
   (* startup initialisation *)
   IF NOT #init OR #T = t#0s THEN
     #init := TRUE;
     #out := #K * #in;
   ELSE
     #out := #out + (#in * #K - #out) * DINT_TO_REAL(DWORD_TO_DINT(#tx) - DWORD_TO_DINT(#last)) / DINT_TO_REAL(T_CONV(#T)) * 1.0E-3;
     IF ABS(#out) < 1.0E-20 THEN #out := 0.0; END_IF;
   END_IF;
   #last := #tx;


   (*
   hm 1.1.2007 rev 1.1
     corrected error while startup value was not correct
     for very small time values real output would run out of range.

   hm 3.1.2007 rev 1.2
     corrected an error for falling edge failures.
     added output faktor K.

   hm 27. 2. 2007 rev 1.3
     output will be input during init for definitive startup condition.

   hm  15.9.2007 rev 1.4
     changed time() to T_PLC_US() for compatibilitxy resons
     increased internal accuracy to Microseconds instead of Milliseconds

   hm  23. oct 2007  rev 1.5
     added out := in to the init statements

   hm  30. nov 2007  rev 1.6
     changed out to be K * in during initialization

   hm  5. jan 2008 rev 1.7
     improved code for better performance

   hm  16. mar. 2008 rev 1.8
     added type conversion to avoid warning under codesys 3.0

   hm  14. jun. 2008 rev 1.9
     improved code

   hm  11. mar. 2009 rev 1.10
     real constants updated to new systax using dot

   hm  18. jan. 2011 rev 1.11
     avoid underrun of out
   *)
END_FUNCTION_BLOCK

FUNCTION_BLOCK "FT_PT2"   // FB163, SCL
TITLE = FT_PT2
{ S7_Optimized_Access := 'FALSE' }
AUTHOR : hugo
FAMILY : CTRL
NAME : PT2
VERSION : 1.5
// FT_PT2 is a 2nd grade filter with programmable times T, D and faktor K.
// 
// uses: INTEGRATE [FB237]
//       T_PLC_MS [FC64] 
//       STIME [FB64],IDB_STIME [DB64]
   VAR_INPUT
      in : Real;
      T : Time;
      D : Real;
      K : Real := 1.0e+0;
   END_VAR
   VAR_OUTPUT
      out : Real;
   END_VAR
   VAR
      init : Bool;
      int1 : "INTEGRATE";
      int2 : "INTEGRATE";
      tn : Real;
      I1 : Real;
      I2 : Real;
      tn2 : Real;
   END_VAR
BEGIN


   (* startup initialisation *)
   IF NOT #init OR #T = T#0s THEN
       #init := TRUE;
       #out := #K * #in;
       #I2 := #out;
   ELSE
       #tn := DINT_TO_REAL(T_CONV(#T)) * 1.0E-3;
       #tn2 := #tn * #tn;
       #int1(X := #in * #K / #tn2 - #I1 * 0.5 * #D / #tn - #I2 / #tn2, Y := #I1);
       #int2(X := #I1,Y := #I2);
       #out := #I2;
   END_IF;


   (* revision history

   15.1.2007 hm        rev 1.1
       changed formula to new more acurate formula

   hm 15.9.2007        rev 1.2
       deleted unused code for init system time reading tx 

   hm  30.11.2007  rev 1.3
       changed out to be K * in during initialization
       avoind divide by 0 if tn = 0

   hm  3. nov. 2008    rev 1.4
       optimized code and fixed a problem with init

   hm  11. mar. 2009   rev 1.5
       real constants updated to new systax using dot

   *)
END_FUNCTION_BLOCK

FUNCTION_BLOCK "FT_TN16"   // FB164, SCL
TITLE = FT_TN16
{ S7_Optimized_Access := 'FALSE' }
AUTHOR : hugo
FAMILY : CTRL
NAME : TN16
VERSION : 1.1
// FT_TN16 is delay function, it will delay a signal by a specified time : T and will store 16 values of in before they are put thru to out.
// for higher OR lower resolution please use FT_TN8 OR FT_TN64 instead.
// 
// uses: T_PLC_MS [FC64]
//       STIME [FB64],IDB_STIME [DB64]
   VAR_INPUT
      in : Real;
      T : Time;
   END_VAR
   VAR_OUTPUT
      out : Real;
      trig : Bool;
   END_VAR
   VAR
      length : Int := 16;
      X : Array[0..15] of Real;
      cnt : Int;
      last : Time;
      tx : Time;
      init : Bool;
   END_VAR
BEGIN


     (* read system time *)
     #tx := T_CONV(DWORD_TO_DINT("T_PLC_MS"()));

     #trig := FALSE;
     IF NOT #init THEN
       #X[#cnt] := #in;
       #init := TRUE;
       #last := #tx;
     ELSIF #tx - #last >= #T / #length THEN
       IF #cnt = #length - 1 THEN #cnt := 0; ELSE #cnt := #cnt + 1; END_IF;
       #out := #X[#cnt];
       #X[#cnt] := #in;
       #last := #tx;
       #trig := TRUE;
     END_IF;

   (* revision history
   hm    1. jan 2007    rev 1.0
     original version

   hm    16. sep 2007  rev 1.1
     changes time() to T_plc_ms() for compatibility reasons

   *)
END_FUNCTION_BLOCK

FUNCTION_BLOCK "FT_TN64"   // FB165, SCL
TITLE = FT_TN64
{ S7_Optimized_Access := 'FALSE' }
AUTHOR : hugo
FAMILY : CTRL
NAME : TN64
VERSION : 1.1
// FT_TN64 is delay function, it will delay a signal by a specified time : T and will store 64 values of in before they are put thru to out.
// if lower resolution is needed, pls use FT_TN8 or FT_TN16 instead.
// 
// uses: T_PLC_MS [FC64]
//       STIME [FB64],IDB_STIME [DB64]
   VAR_INPUT
      in : Real;
      T : Time;
   END_VAR
   VAR_OUTPUT
      out : Real;
      trig : Bool;
   END_VAR
   VAR
      length : Int := 64;
      X : Array[0..63] of Real;
      cnt : Int;
      last : Time;
      tx : Time;
      init : Bool;
   END_VAR
BEGIN


     (* read system time *)
     #tx := T_CONV(DWORD_TO_DINT("T_PLC_MS"()));

     #trig := FALSE;
     IF NOT #init THEN
       #X[#cnt] := #in;
       #init := TRUE;
       #last := #tx;
     ELSIF #tx - #last >= #T / #length THEN
       IF #cnt = #length - 1 THEN #cnt := 0; ELSE #cnt := #cnt + 1; END_IF;
       #out := #X[#cnt];
       #X[#cnt] := #in;
       #last := #tx;
       #trig := TRUE;
     END_IF;

   (* revision history
   hm    1. jan 2007    rev 1.0
     original version

   hm    16. sep 2007  rev 1.1
     changes time() to T_plc_ms() for compatibility reasons

   *)
END_FUNCTION_BLOCK

FUNCTION_BLOCK "FT_TN8"   // FB166, SCL
TITLE = FT_TN8
{ S7_Optimized_Access := 'FALSE' }
AUTHOR : hugo
FAMILY : CTRL
NAME : TN8
VERSION : 1.1
// FT_TN8 is delay function, it will delay a signal by a specified time : T and will store 8 values of in before they are put thru to out.
// if higher resolution is needed, pls use FT_TN16 or FT_TN64 instead.
// 
// uses: T_PLC_MS [FC64]
//       STIME [FB64],IDB_STIME [DB64]
   VAR_INPUT
      in : Real;
      T : Time;
   END_VAR
   VAR_OUTPUT
      out : Real;
      trig : Bool;
   END_VAR
   VAR
      length : Int := 8;
      X : Array[0..7] of Real;
      cnt : Int;
      last : Time;
      tx : Time;
      init : Bool;
   END_VAR
BEGIN


     #tx := T_CONV(DWORD_TO_DINT("T_PLC_MS"()));
     #trig := FALSE;
     IF NOT #init THEN
       #X[#cnt] := #in;
       #init := TRUE;
       #last := #tx;
     ELSIF #tx - #last >= #T / #length THEN
       IF #cnt = #length - 1 THEN #cnt := 0; ELSE #cnt := #cnt + 1; END_IF;
       #out := #X[#cnt];
       #X[#cnt] := #in;
       #last := #tx;
       #trig := TRUE;
     END_IF;

   (* revision history
   hm    1. jan 2007    rev 1.0
     original version

   hm    16. sep 2007  rev 1.1
     changes time() to T_plc_ms() for compatibility reasons

   *)
END_FUNCTION_BLOCK

FUNCTION_BLOCK "HYST"   // FB167, SCL
TITLE = HYST
{ S7_Optimized_Access := 'FALSE' }
AUTHOR : hugo
FAMILY : CTRL
NAME : HYST
VERSION : 1.0
// This Hystereses function has two modes:
// 1. if on > off then Q will be switched high when in > on and switched low when in < off.
// 2. if on < off then Q will be switched high when in < on and switched low when in > off.
// the output win will be high when in is between low and high.
   VAR_INPUT
      In : Real;
      ON : Real;
      OFF : Real;
   END_VAR
   VAR_OUTPUT
      Q : Bool;
      win : Bool;
   END_VAR
BEGIN


   IF #ON >= #OFF THEN
       IF #In < #OFF THEN
           #Q := FALSE;
           #win := FALSE;
       ELSIF  #In > #ON THEN
           #Q := TRUE;
           #win := FALSE;
       ELSE
           #win := TRUE;
       END_IF;
   ELSE
       IF #In > #OFF THEN
           #Q := FALSE;
           #win := FALSE;
       ELSIF  #In < #ON THEN
           #Q := TRUE;
           #win := FALSE;
       ELSE
           #win := TRUE;
       END_IF;
   END_IF;


   (* revision history
   hm      2.  jun 2008    rev 1.0
       original version

   *)
END_FUNCTION_BLOCK

FUNCTION_BLOCK "HYST_1"   // FB168, SCL
TITLE = HYST_1
{ S7_Optimized_Access := 'FALSE' }
AUTHOR : hugo
FAMILY : CTRL
NAME : HYST_1
VERSION : 1.1
// this hysteresis function switches the output high if the input signal reaches obove high and will switch to low when the input falls back below low value.
// a separate output mid is set if the input stays between low and high value.
   VAR_INPUT
      In : Real;
      high : Real;
      low : Real;
   END_VAR
   VAR_OUTPUT
      Q : Bool;
      win : Bool;
   END_VAR
BEGIN


   IF #In < #low THEN
       #Q := FALSE;
       #win := FALSE;
   ELSIF #In > #high THEN
       #Q := TRUE;
       #win := FALSE;
   ELSE
       #win := TRUE;
   END_IF;

   (* code used for rev 1.0
   IF Q THEN
       IF in < low THEN q := FALSE; END_IF;
   ELSE
       IF in > high THEN q := TRUE; END_IF;
   END_IF;
   win := in > low AND in < high;
   *)


   (* revision history
   hm      4.  aug. 2006   rev 1.0
       original version

   hm      2. jun. 2008    rev 1.1
       improved performance
   *)
END_FUNCTION_BLOCK

FUNCTION_BLOCK "HYST_2"   // FB169, SCL
TITLE = HYST_2
{ S7_Optimized_Access := 'FALSE' }
AUTHOR : oscat
FAMILY : CTRL
NAME : HYST_2
VERSION : 1.2
// this hysteresis function switches the output high if the input signal reaches obove val + hys/2 and will switch to low when the input falls back below val - hys/2 value.
// a separate output mid is set if the input stays between low and high value.
   VAR_INPUT
      IN : Real;
      VAL : Real;
      HYS : Real;
   END_VAR
   VAR_OUTPUT
      Q : Bool;
      WIN : Bool;
   END_VAR
   VAR
      tmp : Real;
   END_VAR
BEGIN


   #tmp := #VAL - #HYS * 0.5;
   IF #IN < #tmp THEN
       #Q := FALSE;
       #WIN := FALSE;
   ELSIF #IN > #tmp + #HYS THEN
       #Q := TRUE;
       #WIN := FALSE;
   ELSE
       #WIN := TRUE;
   END_IF;

   (* code used for 1.2 and before
   X := hys * 0.5;
   IF Q THEN
       IF in < val - x THEN q := FALSE; END_IF;
   ELSE
       IF in > val + x THEN q := TRUE; END_IF;
   END_IF;
   win := in > val - x AND in < val + x;
   *)

   (* revision history
   hm      4. aug 2006 rev 1.0
       original version

   hm      5. jan 2008 rev 1.1
       improved code for better performance

   hm      2. jun. 2008    rev 1.2
       improved performance
   *)
END_FUNCTION_BLOCK

FUNCTION_BLOCK "HYST_3"   // FB170, SCL
TITLE = HYST_3
{ S7_Optimized_Access := 'FALSE' }
AUTHOR : oscat
FAMILY : CTRL
NAME : HYST_3
VERSION : 1.2
// this is a double hysteresis function. Out1 follows a hysteresis function defined by val1and hyst, while out 2 follows val2 and hyst.
// if the input signal is between the two hysteresis switches (val1 and val2) then non of the outputs is active.
   VAR_INPUT
      in : Real;
      hyst : Real;
      val1 : Real;
      val2 : Real;
   END_VAR
   VAR_OUTPUT
      Q1 : Bool;
      Q2 : Bool;
   END_VAR
   VAR
      X : Real;
   END_VAR
BEGIN


     #X := #hyst * 0.5;

     IF #in < #val1 - #X THEN
         #Q1 := TRUE;
     ELSIF #in > #val1 + #X THEN
         #Q1 := FALSE;
     END_IF;
     IF #in < #val2 - #X THEN
         #Q2 := FALSE;
     ELSIF #in > #val2 + #X THEN
         #Q2 := TRUE;
     END_IF;

   (* revision history
   hm  22. jan 2007  rev 1.0
     original version

   hm  27. dec 2007  rev 1.1
     changed code for better performance

   hm  5. jan 2008   rev 1.2
     further performance iprovements

   *)
END_FUNCTION_BLOCK

FUNCTION_BLOCK "INTEGRATE"   // FB237, SCL
TITLE = INTEGRATE
{ S7_Optimized_Access := 'FALSE' }
AUTHOR : hugo
FAMILY : CTRL
NAME : INTEGR
VERSION : 1.0
// integrate is a plain integrator with I/O for out.
// 
// uses: T_PLC_MS [FC64]
//       STIME [FB64],IDB_STIME [DB64]
   VAR_INPUT
      "E" : Bool := TRUE;
      X : Real;
      K : Real := 1.0e+0;
   END_VAR
   VAR_IN_OUT
      Y : Real;
   END_VAR
   VAR
      X_last : Real;
      init : Bool;
      last : DWord;
      tx : DWord;
   END_VAR
   VAR_TEMP
      TOP_SI : Struct
         EV_CLASS : Byte;
         EV_NUM : Byte;
         PRIORITY : Byte;
         NUM : Byte;
         TYP2_3 : Byte;
         TYP1 : Byte;
         ZI1 : Word;
         ZI2_3 : DWord;
      END_STRUCT;
      START_UP_SI : Struct
         EV_CLASS : Byte;
         EV_NUM : Byte;
         PRIORITY : Byte;
         NUM : Byte;
         TYP2_3 : Byte;
         TYP1 : Byte;
         ZI1 : Word;
         ZI2_3 : DWord;
      END_STRUCT;
      ERR : Int;
   END_VAR
BEGIN


   (* read actual startup info *)
   (* OB1_SCAN_1  BYTE  -  B#16#01: Abschluss des Neustarts (Warmstarts)
                        -  B#16#02: Abschluss des Wiederanlaufs
                        -  B#16#03: Abschluss des freien Zyklus
                        -  B#16#04: Abschluss des Kaltstarts
                        -  B#16#05: Erster OB 1-Zyklus der neuen Master-CPU nach 
                                    Master-Reserve-Umschaltung und STOP des 
                                    bisherigen Masters *)

   #ERR := RD_SINFO (TOP_SI => #TOP_SI, START_UP_SI => #START_UP_SI);

   (* reset last_time on system startup *)
   IF #TOP_SI.EV_NUM = 1 OR #TOP_SI.EV_NUM = 2 OR #TOP_SI.EV_NUM = 4 THEN 
       #init := FALSE;
   END_IF;

   (*read system time *)
   #tx := "T_PLC_MS"();

   IF NOT #init THEN
       #init := TRUE;
       #X_last := #X;
   ELSIF #"E" THEN
       #Y := (#X + #X_last) * 0.5E-3 * DINT_TO_REAL(DWORD_TO_DINT(#tx)-DWORD_TO_DINT(#last)) * #K + #Y;
       #X_last := #X;
   END_IF;
   #last := #tx;


   (*
   hm  3. nov. 2008    rev 1.0
   original version

   *)
END_FUNCTION_BLOCK

FUNCTION "T_PLC_MS" : DWord   // FC64, SCL
TITLE = T_PLC_MS
{ S7_Optimized_Access := 'FALSE' }
AUTHOR : hugo
FAMILY : MEASURE
NAME : T_PLC_MS
VERSION : 1.2
// T_PLC_MS reads the internal PLC timer and return the time, it has the advantage to be able to set a debug mode 
// and speed up the counter to test the plc timer overrun which occurs every 50 days respectively 25 days at siemens S7
// this routine also allows to correct the behavior of s7 where the internal plc counter will not count all 32 bits.
// 
// uses: STIME [FB64],IDB_STIME [DB64]
BEGIN


   "IDB_STIME"(); 
   #T_PLC_MS := "IDB_STIME".tx; 
   (* hier muss die korrektur für step7 stattfinden
   plctime muss den vollen wertebereich von time ausnutzen:
   wenn bei step7 time -24tage bis plus 24 tage ist dann muss der timer auch beim überlauf auf -24tage springen 
   und auf keinen fall auf 0 !!!!
   für siemens muss ein weiterer fb im main eingebunden werden der sicherstellt das alle 32 bits durchgezählt werden.
   es kann nur ein fb sein den er muss sich das oberste (32te) bit merken.
   oder etwa spring s7 bei überlauf auf -24 tage????? dann wäre keine korrektur nötig.
   *)
   IF "debug" THEN
       #T_PLC_MS := DINT_TO_DWORD((DWORD_TO_DINT(SHL(IN:=#T_PLC_MS,N:="N") OR SHL(IN:=DWORD#1,N:="N"))-1) + DWORD_TO_DINT("offset_1"));
   END_IF;


   (* revision history
   hm  14.9.2007   rev 1.0
       original version

   hm  12. nov 2007    rev 1.1
       added temporaray variable tx because some compilers could not handle time() as an argument

   hm  16. nov. 2008   rev 1.2
       initialized constants with 0 for compatibility reasons
   *)
END_FUNCTION

FUNCTION "T_PLC_US" : DWord   // FC65, SCL
TITLE = T_PLC_US
{ S7_Optimized_Access := 'FALSE' }
AUTHOR : hugo
FAMILY : MEASURE
NAME : T_PLC_US
VERSION : 1.2
// T_PLC_US reads the internal PLC timer and return the time, it has the advantage to be able to set a debug mode 
// and speed up the counter to test the plc timer overrun which occurs every 50 days respectively 25 days at siemens S7
// this routine also allows to correct the behavior of s7 where the internal plc counter will not count all 32 bits.
// 
// uses: STIME [FB64],IDB_STIME [DB64]
BEGIN


   "IDB_STIME"(); 
   #T_PLC_US := DINT_TO_DWORD(DWORD_TO_DINT("IDB_STIME".tx) * 1000); 
   (* hier muss die korrektur für step7 stattfinden
   plctime muss den vollen wertebereich von time ausnutzen:
   wenn bei step7 time -24tage bis plus 24 tage ist dann muss der timer auch beim überlauf auf -24tage springen 
   und auf keinen fall auf 0 !!!!
   für siemens muss ein weiterer fb im main eingebunden werden der sicherstellt das alle 32 bits durchgezählt werden.
   es kann nur ein fb sein den er muss sich das oberste (32te) bit merken.
   oder etwa spring s7 bei überlauf auf -24 tage????? dann wäre keine korrektur nötig.
   *)
   IF "debug" THEN
       #T_PLC_US := DINT_TO_DWORD((DWORD_TO_DINT(SHL(IN:=#T_PLC_US,N:="N") OR SHL(IN:=DWORD#1,N:="N"))-1) + DWORD_TO_DINT("offset_1"));
   END_IF;


   (* revision history
   hm  14.9.2007   rev 1.0
       original version

   hm  12. nov 2007    rev 1.1
       added temporaray variable tx because some compilers could not handle time() as an argument

   hm  16. nov. 2008   rev 1.2
       initialized constants with 0 for compatibility reasons

   *)
END_FUNCTION

FUNCTION "R2_ADD" : "REAL2"   // FC144, SCL
TITLE = R2_ADD
{ S7_Optimized_Access := 'FALSE' }
AUTHOR : hugo
FAMILY : R2
NAME : ADD
VERSION : 1.0
// R2_add adds a real to a double real which extends the accuracy of a real to twice as many digits
//  
// uses: REAL2 [UDT11]
   VAR_INPUT
      X : "REAL2";
      Y : Real;
   END_VAR
   VAR_TEMP
      temp : Real;
      tR2_ADD : "REAL2";
   END_VAR
BEGIN


   #temp := #X.RX;
   #tR2_ADD.RX := #Y + #X.R1 + #X.RX;
   #tR2_ADD.R1 := #temp - #tR2_ADD.RX + #Y + #X.R1;

   #R2_ADD := #tR2_ADD;

   (* revision history
   hm      20.3.2008   rev 1.0
       original version

   *)
END_FUNCTION

FUNCTION "R2_SET" : "REAL2"   // FC147, SCL
TITLE = R2_SET
{ S7_Optimized_Access := 'FALSE' }
AUTHOR : hugo
FAMILY : R2
NAME : SET
VERSION : 1.1
// R2_set sets a double precision real to a single real value.
// 
// uses: REAL2 [UDT11]
   VAR_INPUT
      X : Real;
   END_VAR
   VAR_TEMP
      tR2_SET : "REAL2";
   END_VAR
BEGIN


   #tR2_SET.RX := #X;
   #tR2_SET.R1 := 0.0;

   #R2_SET := #tR2_SET;


   (* revision history
   hm  2. jun. 2008    rev 1.0
       original version

   hm  10. mar. 2009   rev 1.1
       real constants updated to new systax using dot

   *)
END_FUNCTION

FUNCTION "MULTIME" : Time   // FC203, SCL
TITLE = MULTIME
{ S7_Optimized_Access := 'FALSE' }
AUTHOR : hugo
FAMILY : TIDT
NAME : MULTIME
VERSION : 1.1
// multiplies a time by a real number and returns a time
   VAR_INPUT
      t : Time;
      "M" : Real;
   END_VAR
BEGIN


     #MULTIME := T_CONV(REAL_TO_DINT(DINT_TO_REAL(T_CONV(#t))*#"M"));

   (* revision history
   hm      2. oct 2006 rev 1.0
       original version

   hm      14. mar 2008    rev 1.1
       rounded the result after the last digit

   *)
END_FUNCTION

FUNCTION "CTRL_IN" : Real   // FC363, SCL
TITLE = CTRL_IN
{ S7_Optimized_Access := 'FALSE' }
AUTHOR : hugo
FAMILY : CTRL
NAME : CTRL_IN
VERSION : 1.0
// uses: DEAD_ZONE [FC365]
   VAR_INPUT
      SET_POINT : Real;
      ACTUAL : Real;
      NOISE : Real;
   END_VAR
BEGIN


   (* calculate the process error DIFF *)
   #CTRL_IN := "DEAD_ZONE"(X:=#SET_POINT - #ACTUAL,L:=#NOISE);


   (* revision history
   hm  2. jun. 2008    rev 1.0
       original version

   *)
END_FUNCTION

FUNCTION "DEAD_BAND" : Real   // FC364, SCL
TITLE = DEAD_BAND
{ S7_Optimized_Access := 'FALSE' }
AUTHOR : hugo
FAMILY : CTRL
NAME : DEADBAND
VERSION : 1.2
// DEAD_BAND ist eine lineare Übertragungsfunktion mit Totzone. Die Funktion verschiebt den positiven Teil der Kurve um +L und den negativen Teil der Kurve um -L.
// DEAD_BAND = X - L wenn X > L)
// DEAD_BAND = X + L wenn X < -L
// DEAD_BAND = 0 wenn Abs(X) <= L
   VAR_INPUT
      X : Real;
      L : Real;
   END_VAR
BEGIN


     IF #X > #L THEN
       #DEAD_BAND := #X - #L;
     ELSIF #X < -#L THEN
       #DEAD_BAND := #X + #L;
     ELSE
       #DEAD_BAND := 0.0;
     END_IF;


   (* revision history
   hm  2. nov. 2007  rev 1.0
     original version

   hm  14. jun. 2008 rev 1.1
     improved performance

   hm  18. jan. 2011 rev 1.2
     assign 0 before return
   *)
END_FUNCTION

FUNCTION "DEAD_ZONE" : Real   // FC365, SCL
TITLE = DEAD_ZONE
{ S7_Optimized_Access := 'FALSE' }
AUTHOR : hugo
FAMILY : CTRL
NAME : DEADZONE
VERSION : 1.2
// dead_zone2 is a linear transfer function which follows a linear function except for x is close to 0.
// Y = X if abs(x) > L otherwise its 0.
   VAR_INPUT
      X : Real;
      L : Real;
   END_VAR
BEGIN


   IF ABS(#X) > #L THEN
       #DEAD_ZONE := #X;
   ELSE
       #DEAD_ZONE := 0.0;
   END_IF;


   (* revision history
   hm  12. feb. 2007   rev 1.0
       original version

   hm  14. jun. 2008   rev 1.1
       improved performance

   hm  11. mar. 2009   rev 1.2
       real constants updated to new systax using dot

   *)
END_FUNCTION

FUNCTION "BAND_B" : Byte   // FC410, SCL
TITLE = BAND_B
{ S7_Optimized_Access := 'FALSE' }
AUTHOR : hugo
FAMILY : CTRL
NAME : BAND_B
VERSION : 1.0
// BAND_B will limit X to B <= X <= 255-B. while X < B the resulkt will be 0 and while X > 255-B the output will be 255
// otherwise the result = X.
   VAR_INPUT
      X : Byte;
      "B" : Byte;
   END_VAR
BEGIN


   IF BYTE_TO_INT(#X) < BYTE_TO_INT(#"B") THEN
       #BAND_B := 0;
   ELSIF BYTE_TO_INT(#X) > BYTE_TO_INT(BYTE#255) - BYTE_TO_INT(#"B") THEN
       #BAND_B := 255;
   ELSE
       #BAND_B := #X;
   END_IF;



   (* revision history
   hm  21. nov. 2008   rev 1.0
       original version

   *)
END_FUNCTION

// ===== PLC "Engineering conversion"  Unspecific CPU S7 300 =====

VAR_GLOBAL CONSTANT   // PLC tag table "STEP7 classic symbols"
   "#T0" : Real := -2.731500E+002;   // MigChange: -273.15 OriginalComment: absoluter Nullpunkt in °C
   "PI2" : Real := 6.28318530717958647692528676655900576;   // PI * 2
END_VAR

DATA_BLOCK "LANGUAGE"   // DB4
TITLE = LANGUAGE
{ S7_Optimized_Access := 'FALSE' }
AUTHOR : oscat
FAMILY : CONSTANT
NAME : DBLANG
VERSION : 1.2
   VAR
      DEFAULT : Int := 1;   // 1=english, 2=german, 3=french
      LMAX : Int := 3;
      WEEKDAYS : Array[1..3, 1..7] of String[10];
      WEEKDAYS2 : Array[1..3, 1..7] of String[2];
      MONTHS : Array[1..3, 1..12] of String[10];
      MONTHS3 : Array[1..3, 1..12] of String[3];
      DIRS : Array[1..3, 0..15] of String[3];
   END_VAR
BEGIN
   WEEKDAYS[1,1] := 'Monday';
   WEEKDAYS[1,2] := 'Tuesday';
   WEEKDAYS[1,3] := 'Wednesday';
   WEEKDAYS[1,4] := 'Thursday';
   WEEKDAYS[1,5] := 'Friday';
   WEEKDAYS[1,6] := 'Saturday';
   WEEKDAYS[1,7] := 'Sunday';
   WEEKDAYS[2,1] := 'Montag';
   WEEKDAYS[2,2] := 'Dienstag';
   WEEKDAYS[2,3] := 'Mittwoch';
   WEEKDAYS[2,4] := 'Donnerstag';
   WEEKDAYS[2,5] := 'Freitag';
   WEEKDAYS[2,6] := 'Samstag';
   WEEKDAYS[2,7] := 'Sonntag';
   WEEKDAYS[3,1] := 'Lundi';
   WEEKDAYS[3,2] := 'Mardi';
   WEEKDAYS[3,3] := 'Mercredi';
   WEEKDAYS[3,4] := 'Jeudi';
   WEEKDAYS[3,5] := 'Vendredi';
   WEEKDAYS[3,6] := 'Samedi';
   WEEKDAYS[3,7] := 'Dimanche';
   WEEKDAYS2[1,1] := 'Mo';
   WEEKDAYS2[1,2] := 'Tu';
   WEEKDAYS2[1,3] := 'We';
   WEEKDAYS2[1,4] := 'Th';
   WEEKDAYS2[1,5] := 'Fr';
   WEEKDAYS2[1,6] := 'Sa';
   WEEKDAYS2[1,7] := 'Su';
   WEEKDAYS2[2,1] := 'Mo';
   WEEKDAYS2[2,2] := 'Di';
   WEEKDAYS2[2,3] := 'Mi';
   WEEKDAYS2[2,4] := 'Do';
   WEEKDAYS2[2,5] := 'Fr';
   WEEKDAYS2[2,6] := 'Sa';
   WEEKDAYS2[2,7] := 'So';
   WEEKDAYS2[3,1] := 'Lu';
   WEEKDAYS2[3,2] := 'Ma';
   WEEKDAYS2[3,3] := 'Me';
   WEEKDAYS2[3,4] := 'Je';
   WEEKDAYS2[3,5] := 'Ve';
   WEEKDAYS2[3,6] := 'Sa';
   WEEKDAYS2[3,7] := 'Di';
   MONTHS[1,1] := 'January';
   MONTHS[1,2] := 'February';
   MONTHS[1,3] := 'March';
   MONTHS[1,4] := 'April';
   MONTHS[1,5] := 'May';
   MONTHS[1,6] := 'June';
   MONTHS[1,7] := 'July';
   MONTHS[1,8] := 'August';
   MONTHS[1,9] := 'September';
   MONTHS[1,10] := 'October';
   MONTHS[1,11] := 'November';
   MONTHS[1,12] := 'December';
   MONTHS[2,1] := 'Januar';
   MONTHS[2,2] := 'Februar';
   MONTHS[2,3] := 'März';
   MONTHS[2,4] := 'April';
   MONTHS[2,5] := 'Mai';
   MONTHS[2,6] := 'Juni';
   MONTHS[2,7] := 'Juli';
   MONTHS[2,8] := 'August';
   MONTHS[2,9] := 'September';
   MONTHS[2,10] := 'Oktober';
   MONTHS[2,11] := 'November';
   MONTHS[2,12] := 'Dezember';
   MONTHS[3,1] := 'Janvier';
   MONTHS[3,2] := 'Février';
   MONTHS[3,3] := 'mars';
   MONTHS[3,4] := 'Avril';
   MONTHS[3,5] := 'Mai';
   MONTHS[3,6] := 'Juin';
   MONTHS[3,7] := 'Juillet';
   MONTHS[3,8] := 'Août';
   MONTHS[3,9] := 'Septembre';
   MONTHS[3,10] := 'Octobre';
   MONTHS[3,11] := 'Novembre';
   MONTHS[3,12] := 'Decembre';
   MONTHS3[1,1] := 'Jan';
   MONTHS3[1,2] := 'Feb';
   MONTHS3[1,3] := 'Mar';
   MONTHS3[1,4] := 'Apr';
   MONTHS3[1,5] := 'May';
   MONTHS3[1,6] := 'Jun';
   MONTHS3[1,7] := 'Jul';
   MONTHS3[1,8] := 'Aug';
   MONTHS3[1,9] := 'Sep';
   MONTHS3[1,10] := 'Oct';
   MONTHS3[1,11] := 'Nov';
   MONTHS3[1,12] := 'Dec';
   MONTHS3[2,1] := 'Jan';
   MONTHS3[2,2] := 'Feb';
   MONTHS3[2,3] := 'Mrz';
   MONTHS3[2,4] := 'Apr';
   MONTHS3[2,5] := 'Mai';
   MONTHS3[2,6] := 'Jun';
   MONTHS3[2,7] := 'Jul';
   MONTHS3[2,8] := 'Aug';
   MONTHS3[2,9] := 'Sep';
   MONTHS3[2,10] := 'Okt';
   MONTHS3[2,11] := 'Nov';
   MONTHS3[2,12] := 'Dez';
   MONTHS3[3,1] := 'Jan';
   MONTHS3[3,2] := 'Fev';
   MONTHS3[3,3] := 'Mar';
   MONTHS3[3,4] := 'Avr';
   MONTHS3[3,5] := 'Mai';
   MONTHS3[3,6] := 'Jun';
   MONTHS3[3,7] := 'Jul';
   MONTHS3[3,8] := 'Aou';
   MONTHS3[3,9] := 'Sep';
   MONTHS3[3,10] := 'Oct';
   MONTHS3[3,11] := 'Nov';
   MONTHS3[3,12] := 'Dec';
   DIRS[1,0] := 'N';
   DIRS[1,1] := 'NNE';
   DIRS[1,2] := 'NE';
   DIRS[1,3] := 'ENE';
   DIRS[1,4] := 'E';
   DIRS[1,5] := 'ESE';
   DIRS[1,6] := 'SE';
   DIRS[1,7] := 'SSE';
   DIRS[1,8] := 'S';
   DIRS[1,9] := 'SSW';
   DIRS[1,10] := 'SW';
   DIRS[1,11] := 'WSW';
   DIRS[1,12] := 'W';
   DIRS[1,13] := 'WNW';
   DIRS[1,14] := 'NW';
   DIRS[1,15] := 'NNW';
   DIRS[2,0] := 'N';
   DIRS[2,1] := 'NNO';
   DIRS[2,2] := 'NO';
   DIRS[2,3] := 'ONO';
   DIRS[2,4] := 'O';
   DIRS[2,5] := 'OSO';
   DIRS[2,6] := 'SO';
   DIRS[2,7] := 'SSO';
   DIRS[2,8] := 'S';
   DIRS[2,9] := 'SSW';
   DIRS[2,10] := 'SW';
   DIRS[2,11] := 'WSW';
   DIRS[2,12] := 'W';
   DIRS[2,13] := 'WNW';
   DIRS[2,14] := 'NW';
   DIRS[2,15] := 'NNW';
   DIRS[3,0] := 'N';
   DIRS[3,1] := 'NNO';
   DIRS[3,2] := 'NO';
   DIRS[3,3] := 'ONO';
   DIRS[3,4] := 'O';
   DIRS[3,5] := 'OSO';
   DIRS[3,6] := 'SO';
   DIRS[3,7] := 'SSO';
   DIRS[3,8] := 'S';
   DIRS[3,9] := 'SSW';
   DIRS[3,10] := 'SW';
   DIRS[3,11] := 'WSW';
   DIRS[3,12] := 'W';
   DIRS[3,13] := 'WNW';
   DIRS[3,14] := 'NW';
   DIRS[3,15] := 'NNW';
END_DATA_BLOCK

FUNCTION_BLOCK "ASTRO"   // FB136, SCL
TITLE = ASTRO
{ S7_Optimized_Access := 'FALSE' }
AUTHOR : oscat
FAMILY : CONVERT
NAME : ASTRO
VERSION : 1.1
// this function converts different length units
// any unused input can simply be left open.
// different inputs connected at the same time will be added up.
   VAR_INPUT
      "m" : Real;
      AE : Real;
      PC : Real;
      LJ : Real;
   END_VAR
   VAR_OUTPUT
      Ym : Real;
      YAE : Real;
      YPC : Real;
      YLJ : Real;
   END_VAR
BEGIN


   #YAE :=  #AE
           + #"m" * 6.6845871535E-012
           + #PC * 206265.0
           + #LJ * 63240.0;
   #Ym := #YAE * 149.597870E9;
   #YPC := #YAE * 4.8481322570E-006;
   #YLJ := #YAE * 1.5812776724E-005;


   (*
   Länge Meter m SI-Basiseinheit
   Astronomische Einheit* AE 1 AE = 149,597 870 · E9 m
   Parsec pc 1 pc = 206265 AE = 30,857 · E15 m
   Lichtjahr Lj 1 Lj = 9,460 530 · E15 m = 63240 AE = 0,306 59 pc
   Ångström Å 1 Å = E–l0 m
   typograph. Punkt p 1 p = 0,376 065 mm • im Druckereigewerbe
   inch** in 1 in = 2,54 · E–2 m = 25,4 mm***
   foot ft 1 ft = 0,3048 m = 30,48 cm
   yard yd 1 yd = 0,9144 m
   mile mile 1 mile = 1609,344 m
   Internat. Seemeile sm 1 sm = 1852 m
   Fathom fm 1 fm = 1,829 m • in der Seeschifffahrt
   *)

   (* revision history

   hm  27. mar. 2007   rev 1.0
       original version

   hm  11. mar. 2009   rev 1.1
       improved code

   *)
END_FUNCTION_BLOCK

FUNCTION_BLOCK "ENERGY"   // FB137, SCL
TITLE = ENERGY
{ S7_Optimized_Access := 'FALSE' }
AUTHOR : hugo
FAMILY : CONVERT
NAME : ENERGY
VERSION : 1.2
// this function converts different energy units
// any unused input can simply be left open.
// different inputs connected at the same time will be added up.
   VAR_INPUT
      J : Real;
      C : Real;
      Wh : Real;
   END_VAR
   VAR_OUTPUT
      YJ : Real;
      YC : Real;
      YWh : Real;
   END_VAR
BEGIN


   #YJ := #J + #Wh * 3600.0 + #C * 4.1868;
   #YC := #YJ * 0.238845896627496;
   #YWh := #YJ * 2.7777777778E-004;


   (*
   Arbeit, Energie, Joule* J 1 J = 1 N · m = 1 W · s = (1/3,6) E–6 kW · h = 1 kg · m2/s2
   Wärmemenge Kilowattstunde kW · h 1 kW · h = 3,6 MJ = 860 kcal
   Elektronvolt eV 1 eV = 160,218 92 E–21 J
   Erg erg 1 erg = 1E–7 J
   Kalorie cal 1 cal = 4,1868 J = 1,163 E–3 W · h
   Therm therm 1 therm = 105,50 · 106 J
   *)

   (* revision history

   hm  27. mar. 2007 rev 1.0
     original version

   hm  11. mar. 2009 rev 1.1
     improved code

   hm 16. jan 2010 rev 1.2
     avoid the string cal in comments for codesys import bug


   *)
END_FUNCTION_BLOCK

FUNCTION_BLOCK "LENGTH"   // FB138, SCL
TITLE = LENGTH
{ S7_Optimized_Access := 'FALSE' }
AUTHOR : hugo
FAMILY : CONVERT
NAME : LENGTH
VERSION : 1.1
// this function converts different length units
// any unused input can simply be left open.
// different inputs connected at the same time will be added up.
   VAR_INPUT
      "m" : Real;
      p : Real;
      in : Real;
      ft : Real;
      yd : Real;
      mile : Real;
      sm : Real;
      fm : Real;
   END_VAR
   VAR_OUTPUT
      Ym : Real;
      Yp : Real;
      Yin : Real;
      Yft : Real;
      Yyd : Real;
      Ymile : Real;
      Ysm : Real;
      Yfm : Real;
   END_VAR
BEGIN


   #Ym := #"m"
         + #p * 0.000376065
         + #in * 0.0254
         + #ft * 0.3048
         + #yd * 0.9144
         + #mile * 1609.344
         + #sm * 1852.0
         + #fm * 1.829;
   #Yp := #Ym * 2659.11478068951;
   #Yin := #Ym * 39.37007874016;
   #Yft := #Ym * 3.28083989501;
   #Yyd := #Ym * 1.09361329834;
   #Ymile := #Ym * 0.00062137119;
   #Ysm := #Ym * 0.00053995680;
   #Yfm := #Ym * 0.54674685621;

   (*
   Länge Meter m SI-Basiseinheit
   Astronomische Einheit* AE 1 AE = 149,597 870 · E9 m
   Parsec pc 1 pc = 206265 AE = 30,857 · E15 m
   Lichtjahr Lj 1 Lj = 9,460 530 · E15 m = 63240 AE = 0,306 59 pc
   Ångström Å 1 Å = E–l0 m
   typograph. Punkt p 1 p = 0,376 065 mm • im Druckereigewerbe
   inch** in 1 in = 2,54 · E–2 m = 25,4 mm***
   foot ft 1 ft = 0,3048 m = 30,48 cm
   yard yd 1 yd = 0,9144 m
   mile mile 1 mile = 1609,344 m
   Internat. Seemeile sm 1 sm = 1852 m
   Fathom fm 1 fm = 1,829 m • in der Seeschifffahrt
   *)

   (* revision history

   hm  27. mar. 2007    rev 1.0
       original version

   hm  11. mar. 2009   rev 1.1
       improved code

   *)
END_FUNCTION_BLOCK

FUNCTION_BLOCK "PRESSURE"   // FB139, SCL
TITLE = PRESSURE
{ S7_Optimized_Access := 'FALSE' }
AUTHOR : hugo
FAMILY : CONVERT
NAME : PRESSUR
VERSION : 1.1
// this function converts different pressure units
// any unused input can simply be left open.
// different inputs connected at the same time will be added up.
   VAR_INPUT
      mws : Real;
      torr : Real;
      att : Real;
      atm : Real;
      pa : Real;
      bar : Real;
   END_VAR
   VAR_OUTPUT
      Ymws : Real;
      Ytorr : Real;
      Yatt : Real;
      Yatm : Real;
      Ypa : Real;
      Ybar : Real;
   END_VAR
BEGIN


   #Ybar := #bar +
         #pa / 1.0E-5 +
         0.980665 * #att +
         1.01325 * #atm +
         0.001333224 * #torr +
         0.0980665 * #mws;
   #Ymws := #Ybar * 10.1971621297793;
   #Ytorr := #Ybar * 750.0615050434140;
   #Yatt := #Ybar * 1.0197162129779;
   #Yatm := #Ybar * 0.9869232667160;
   #Ypa := #Ybar * 100000.0;


   (*
   Druck, Pascal Pa 1 Pa = 1 N/m2 = 1 kg/(s2 E m) . 0,75 E 10.2 mmHg
   mechanische 1 MPa = 1 N/mm2 . fur Festigkeitsangaben
   Spannung Bar bar 1 bar = 105 Pa = 103 mbar = 105 kg/(s2 E m)
   Millimeter- mmHg 1 mmHg = 133,322 Pa = 1,333 22 mbar
   Quecksilbersaule . nur in Heilkunde zulassig
   physik. Atmosphare atm 1 atm = 1,013 25 bar
   techn. Atmosphare at 1 at = 1 kp/cm2 = 0,980665 bar
   Torr Torr 1 Torr = (101325/760) Pa = 1,333224 mbar
   Meter-Wassersaule mWS 1 mWS = 9806,65 Pa = 98,0665 mbar
   psi lbf/in2 1 lbf/in2 = 68,947 57 mbar = 6894,757 Pa

   *)

   (* revision history

   hm  27. mar. 2007   rev 1.0
       original version

   hm  11. mar. 2009 rev 1.1
       improved code

   *)
END_FUNCTION_BLOCK

FUNCTION_BLOCK "SPEED"   // FB140, SCL
TITLE = SPEED
{ S7_Optimized_Access := 'FALSE' }
AUTHOR : hugo
FAMILY : CONVERT
NAME : SPEED
VERSION : 1.1
// this function converts different speed units
// any unused input can simply be left open.
// different inputs connected at the same time will be added up.
   VAR_INPUT
      ms : Real;
      kmh : Real;
      kn : Real;
      mh : Real;
   END_VAR
   VAR_OUTPUT
      Yms : Real;
      Ykmh : Real;
      Ykn : Real;
      Ymh : Real;
   END_VAR
BEGIN


   #Yms := #ms +
           #kmh * 0.27777777777778 +
           #kn * 0.5144444 +
           #mh * 0.44704;
   #Ykmh := #Yms * 3.6;
   #Ykn := #Yms * 1.94384466037535;
   #Ymh := #Yms * 2.23693629205440;


   (*
   Geschwindigkeit Meter durch Sekunde m/s 1 m/s = 3,6 km/h
   km durch (pro) Stunde, nicht „Stundenkilometer“ verwenden
   Knoten kn 1 kn = 1 sm/h = 0,5144 m/s

   *)

   (* revision history
   hm  27. mar. 2009   rev 1.0
       original version

   hm  11. mar. 2009   rev 1.1
       improved code

   *)
END_FUNCTION_BLOCK

FUNCTION_BLOCK "TEMPERATURE"   // FB141, SCL
TITLE = TEMPERATURE
{ S7_Optimized_Access := 'FALSE' }
AUTHOR : hugo
FAMILY : CONVERT
NAME : TEMP
VERSION : 1.0
// this function converts different temperature units
// any unused input can simply be left open.
// different inputs connected at the same time will be added up.
   VAR_INPUT
      K : Real;
      C : Real := -2.7315e+2;
      F : Real := -4.5967e+2;
      Re : Real := -2.1852e+2;
      Ra : Real;
   END_VAR
   VAR_OUTPUT
      YK : Real;
      YC : Real;
      YF : Real;
      YRe : Real;
      YRa : Real;
   END_VAR
BEGIN


     #YK := #K + (#C + 273.15) + (#F + 459.67) * 0.555555555555 + (#Re * 1.25 + 273.15) + (#Ra * 0.555555555555);
     #YC := #YK -273.15;
     #YF := #YK * 1.8 - 459.67;
     #YRe := (#YK - 273.15) * 0.8;
     #YRa := #YK * 1.8;


   (* revision history
   hm  21. feb. 2008 rev 1.0
     original version

   *)
END_FUNCTION_BLOCK

FUNCTION "BFT_TO_MS" : Real   // FC349, SCL
TITLE = BFT_TO_MS
{ S7_Optimized_Access := 'FALSE' }
AUTHOR : hugo
FAMILY : CONVERT
NAME : BFT2MS
VERSION : 1.0
// this function converts wind speed from beaufort to m/s
   VAR_INPUT
      BFT : Int;
   END_VAR
BEGIN


     #BFT_TO_MS := (#BFT**1.5) * 0.836;


   (* revision history
   hm  12. 6. 2008     rev 1.0
       original version

   *)
END_FUNCTION

FUNCTION "C_TO_F" : Real   // FC350, SCL
TITLE = C_TO_F
{ S7_Optimized_Access := 'FALSE' }
AUTHOR : hugo
FAMILY : CONVERT
NAME : C2F
VERSION : 1.1
// this function converts celsius  to fahrenheit
   VAR_INPUT
      celsius : Real;
   END_VAR
BEGIN


   #C_TO_F := #celsius * 1.8 + 32.0;


   (* revision history

   hm  4. aug. 2006    rev 1.0
       original version

   hm  11. mar. 2009   rev 1.1
       real constants updated to new systax using dot

   *)
END_FUNCTION

FUNCTION "C_TO_K" : Real   // FC351, SCL
TITLE = C_TO_K
{ S7_Optimized_Access := 'FALSE' }
AUTHOR : hugo
FAMILY : CONVERT
NAME : C2K
VERSION : 1.1
// this function converts celsius to kelvin
   VAR_INPUT
      Celsius : Real;
   END_VAR
BEGIN


     #C_TO_K := #Celsius - "#T0";


   (* revision history

   hm 4. aug 2006 rev 1.0
    original version

   hm 19. aug 2009 rev 1.1
    fixed calculation error

   *)
END_FUNCTION

FUNCTION "DEG_TO_DIR" : String[254]   // FC352, SCL
TITLE = DEG_TO_DIR
{ S7_Optimized_Access := 'FALSE' }
AUTHOR : hugo
FAMILY : CONVERT
NAME : DEG2DIR
VERSION : 1.1
// this function converts degrees in compass direction.
// the function supports output in english (L=0) and german (L=1).
// 
// uses: LANGUAGE [DB4]
   VAR_INPUT
      DEG : Int;
      N : Int;
      L : Int;
   END_VAR
   VAR_TEMP
      tDEG_TO_DIR : String[3];
      ly : Int;
   END_VAR
BEGIN


   #tDEG_TO_DIR := #DEG_TO_DIR;

   IF #L = 0 THEN 
       #ly := "LANGUAGE".DEFAULT; 
   ELSE 
       #ly := MIN(IN1:=#L, IN2:="LANGUAGE".LMAX); 
   END_IF;
   #DEG_TO_DIR := "LANGUAGE".DIRS[#ly, ((WORD_TO_INT(SHL(IN:=INT_TO_WORD(#DEG),N:=#N-1)) + 45) / 90) MOD WORD_TO_INT(SHL(IN:=WORD#0002,N:=#N))*WORD_TO_INT(SHR(IN:=WORD#0008,N:=#N))];

   #DEG_TO_DIR := #tDEG_TO_DIR;

   (*
   DIR := ((SHL(DEG,N-1) + 45) / 90) MOD SHL(INT#2,N);
   explanation :
   DIR is calculated BY the following formula:
   DIR := ((DIR + 45) / 90) MOD 4 if N = 1 digit
   North = 0, East = 1 ....
   DIR := ((DIR + 22,5) / 45) MOD 8 if N = 2 digit
   convert to integer calculation
   DIR := ((DIR*2 + 45) / 90) MOD 8
   N = 0, NE = 1 ....
   ther above formula replaces 2^N with shift for performance
   *)



   (* revision histroy
   hm  11. jun. 2008   rev 1.0
       original release

   hm  22. oct. 2008   rev 1.1
       changed size of string variables to 30
   *)
END_FUNCTION

FUNCTION "DIR_TO_DEG" : Int   // FC353, SCL
TITLE = DIR_TO_DEG
{ S7_Optimized_Access := 'FALSE' }
AUTHOR : hugo
FAMILY : CONVERT
NAME : DIR2DEG
VERSION : 1.1
// this function converts compass directions to degrees
// it will recognize up to 3 letter directions in english and german writing.
// 
// uses: LANGUAGE [DB4]
//       EQ_STRNG [FC10]
   VAR_INPUT
      DIR : String[254];
      L : Int;
   END_VAR
   VAR_TEMP
      ly : Int;
      i : Int;
      tDIR : String[3];
   END_VAR
BEGIN


   #tDIR := #DIR;

   IF #L = 0 THEN #ly := "LANGUAGE".DEFAULT; ELSE #ly := MIN(IN1:=#L, IN2:="LANGUAGE".LMAX); END_IF;
   FOR #i := 0 TO 15 DO
       IF "LANGUAGE".DIRS[#ly, #i] S_COMP #tDIR THEN EXIT; END_IF;
   END_FOR;
   #DIR_TO_DEG := WORD_TO_INT(SHR(IN:=INT_TO_WORD(#i * 45 + 1), N:=1));

   (* revision histroy
   hm  22. oct. 2008   rev 1.1
       original release

   *)
END_FUNCTION

FUNCTION "F_TO_C" : Real   // FC354, SCL
TITLE = F_TO_C
{ S7_Optimized_Access := 'FALSE' }
AUTHOR : hugo
FAMILY : CONVERT
NAME : F2C
VERSION : 1.1
// this FUNCTION converts fahrenheit TO celsius
   VAR_INPUT
      fahrenheit : Real;
   END_VAR
BEGIN


   #F_TO_C := (#fahrenheit - 32.0) * 0.5555555555555;


   (* revision history
   hm  4. aug 2006 rev 1.0
       original version

   hm  11. mar. 2009   rev 1.1
       real constants updated to new systax using dot

   *)
END_FUNCTION

FUNCTION "F_TO_OM" : Real   // FC355, SCL
TITLE = F_TO_OM
{ S7_Optimized_Access := 'FALSE' }
AUTHOR : hugo
FAMILY : CONVERT
NAME : F2OM
VERSION : 1.1
// this function converts frequency to Omega F
// Omega = 2*PI*F
   VAR_INPUT
      F : Real;
   END_VAR
BEGIN


   #F_TO_OM := "PI2" * #F;

   (*  Käse!
       F_TO_OM := math.PI2 * F;
   *)

   (* revision history
   hm  22. jan. 2007   rev 1.0
       original version

   hm  18. oct. 2008   rev 1.1
       unsing math constants

   *)
END_FUNCTION

FUNCTION "F_TO_PT" : Time   // FC356, SCL
TITLE = F_TO_PT
{ S7_Optimized_Access := 'FALSE' }
AUTHOR : hugo
FAMILY : CONVERT
NAME : F2PT
VERSION : 1.1
// this function converts frequency to periode time
   VAR_INPUT
      F : Real;
   END_VAR
BEGIN


   #F_TO_PT := T_CONV(REAL_TO_DINT(1.0 / #F * 1000.0));


   (* revision history

   hm  4. aug. 2006    rev 1.0
       original version

   hm  11. mar. 2009   rev 1.1
       real constants updated to new systax using dot

   *)
END_FUNCTION

FUNCTION "KMH_TO_MS" : Real   // FC357, SCL
TITLE = KMH_TO_MS
{ S7_Optimized_Access := 'FALSE' }
AUTHOR : hugo
FAMILY : CONVERT
NAME : KMH2MS
VERSION : 1.1
// this function converts velocities from Kilometers / hour to Meters / Second
   VAR_INPUT
      kmh : Real;
   END_VAR
BEGIN


     #KMH_TO_MS := #kmh * 0.2777777777777;

   (* revision history
   hm  4. feb 2007   rev 1.0
     original version

   hm  6. jan 2008   rev 1.1
     improved performance

   *)
END_FUNCTION

FUNCTION "MS_TO_BFT" : Int   // FC358, SCL
TITLE = MS_TO_BFT
{ S7_Optimized_Access := 'FALSE' }
AUTHOR : hugo
FAMILY : CONVERT
NAME : MS2BFT
VERSION : 1.0
// this function converts wind speed from M/s to beaufort
   VAR_INPUT
      MS : Real;
   END_VAR
BEGIN


   #MS_TO_BFT := REAL_TO_INT((#MS * 1.196172)**0.666667);


   (* revision history
   hm  12. 6. 2008     rev 1.0
       original version

   *)
END_FUNCTION

FUNCTION "MS_TO_KMH" : Real   // FC359, SCL
TITLE = MS_TO_KMH
{ S7_Optimized_Access := 'FALSE' }
AUTHOR : hugo
FAMILY : CONVERT
NAME : MS2KMH
VERSION : 1.0
// this function converts velocities from Meters / Second to Kilometers / hour.
   VAR_INPUT
      ms : Real;
   END_VAR
BEGIN


     #MS_TO_KMH := #ms * 3.6;
END_FUNCTION

FUNCTION "K_TO_C" : Real   // FC360, SCL
TITLE = K_TO_C
{ S7_Optimized_Access := 'FALSE' }
AUTHOR : hugo
FAMILY : CONVERT
NAME : K2C
VERSION : 1.1
// this function converts kelvin to celsius
   VAR_INPUT
      Kelvin : Real;
   END_VAR
BEGIN


     #K_TO_C := #Kelvin + "#T0";


   (* revision history

   hm 4. aug 2006 rev 1.0
    original version

   hm 19. aug 2009 rev 1.1
    fixed calculation error

   *)
END_FUNCTION

FUNCTION "OM_TO_F" : Real   // FC361, SCL
TITLE = OM_TO_F
{ S7_Optimized_Access := 'FALSE' }
AUTHOR : hugo
FAMILY : CONVERT
NAME : OM2F
VERSION : 1.1
// this function converts Omega F to frequency
// F = OM / (2*PI)
   VAR_INPUT
      OM : Real;
   END_VAR
BEGIN


   #OM_TO_F := #OM / "PI2";

   (*  Käse!
       OM_TO_F := OM / math.PI2;
   *)

   (* revision history
   hm  22. jan. 2007   rev 1.0
       original version

   hm  18. oct. 2008   rev 1.1
       using math constants

   *)
END_FUNCTION

FUNCTION "PT_TO_F" : Real   // FC362, SCL
TITLE = PT_TO_F
{ S7_Optimized_Access := 'FALSE' }
AUTHOR : hugo
FAMILY : CONVERT
NAME : PT2F
VERSION : 1.1
// this function converts periode time to frequency
   VAR_INPUT
      PT : Time;
   END_VAR
BEGIN


   #PT_TO_F := 1000.0 / DINT_TO_REAL(T_CONV(#PT));


   (*  revision history
   hm  4. aug. 2006    rev 1.0
       original version

   hm  11. mar. 2009   rev 1.1
       real constants updated to new systax using dot

   *)
END_FUNCTION

FUNCTION "GEO_TO_DEG" : Real   // FC413, SCL
TITLE = GEO_TO_DEG
{ S7_Optimized_Access := 'FALSE' }
AUTHOR : hugo
FAMILY : CONVERT
NAME : GEO2DEG
VERSION : 1.0
// this function converts degrees, minutes seconds to decimal degrees.
   VAR_INPUT
      D : Int;
      "M" : Int;
      SEC : Real;
   END_VAR
BEGIN


   #GEO_TO_DEG := INT_TO_REAL(#D) + INT_TO_REAL(#"M") * 0.016666666666667 + #SEC * 0.00027777777777778;

   (* revision histroy
   hm  22. jan. 2009    rev 1.0
       original release


   *)
END_FUNCTION

// ===== PLC "Engineering measurements"  Unspecific CPU S7 300 =====

VAR_GLOBAL CONSTANT   // PLC tag table "STEP7 classic symbols"
   "debug" : Bool := FALSE;
   "N" : Int := 0;
   "offset" : Int := 0;
   "offset_1" : DWord := 0;
END_VAR

TYPE "REAL2"
VERSION : 0.0
   STRUCT
      R1 : Real;
      RX : Real;
   END_STRUCT;
END_TYPE

DATA_BLOCK "IDB_STIME"   // DB64
{ S7_Optimized_Access := 'FALSE' }
AUTHOR : dalbi
FAMILY : MEASURE
VERSION : 0.0
// stored: InstanceOfName STIME
"STIME"
BEGIN
END_DATA_BLOCK

FUNCTION_BLOCK "STIME"   // FB64, SCL
TITLE = STIME
{ S7_Optimized_Access := 'FALSE' }
AUTHOR : dalbi
FAMILY : MEASURE
NAME : STIME
VERSION : 1.4
// this function block makes sure that the timer of a siemens sps counts from 0 - 2^32-1.
   VAR_OUTPUT
      tx : DWord;
      at_tx AT tx : Array[0..31] of Bool;
   END_VAR
   VAR
      last_time : DWord;
      bit31 : Bool;
      init : Bool := TRUE;
   END_VAR
   VAR_TEMP
      TOP_SI : Struct
         EV_CLASS : Byte;
         EV_NUM : Byte;
         PRIORITY : Byte;
         NUM : Byte;
         TYP2_3 : Byte;
         TYP1 : Byte;
         ZI1 : Word;
         ZI2_3 : DWord;
      END_STRUCT;
      START_UP_SI : Struct
         EV_CLASS : Byte;
         EV_NUM : Byte;
         PRIORITY : Byte;
         NUM : Byte;
         TYP2_3 : Byte;
         TYP1 : Byte;
         ZI1 : Word;
         ZI2_3 : DWord;
      END_STRUCT;
      ERR : Int;
   END_VAR
BEGIN


   (* this FB is only necessary for siemens sps
   the siemens sps timer counts from 0 to 2^31-1 and starts at 0 sfter overrun.
   this means that the bit 31 (the highest bit ) will never be used and therefore
   a problem arises when t2 - t1 is checked.
   t2 - t1 is always valid also in an timer overrun situation where the time t1 is very high and t2 is very low.
   the result of the subtraction t2 - t1 however is still valid.
   this calculation does not work for soiemens because the highest bit is not used.

   this module stores the highest bit, changes the highest bit at every overrun occurence and stuffs ther highest bit in the output.
   the output is then used by t_plc_us and t_plc_ms.

   the correction needs and fb and not a function because the value of the highest bit has to be stored.

   do never use this function block in a codesys environment. the timer in codesys is correct and runs from 0 to 2^32-1
   *)

   (* read actual startup info *)
   (* OB1_SCAN_1  BYTE  -  B#16#01: Abschluss des Neustarts (Warmstarts)
                        -  B#16#02: Abschluss des Wiederanlaufs
                        -  B#16#03: Abschluss des freien Zyklus
                        -  B#16#04: Abschluss des Kaltstarts
                        -  B#16#05: Erster OB 1-Zyklus der neuen Master-CPU nach 
                                    Master-Reserve-Umschaltung und STOP des 
                                    bisherigen Masters *)

   #ERR := RD_SINFO (TOP_SI => #TOP_SI, START_UP_SI => #START_UP_SI);

   (* reset last_time on system startup *)
   IF #TOP_SI.EV_NUM = 1 OR #TOP_SI.EV_NUM = 2 OR #TOP_SI.EV_NUM = 4 OR NOT #init THEN 
       #last_time := 0;
       #bit31 := false;
       #init := true;
   END_IF;

   (* read the system timer *)
   #tx := DINT_TO_DWORD(T_CONV(TIME_TCK()));

   (* check for overrun *)
   IF DWORD_TO_DINT(#tx) < DWORD_TO_DINT(#last_time) THEN
       (* an overrun has occured, change the value of the highest bit *)
       #bit31 := NOT #bit31;
   END_IF;

   (* stuff the highest bit into the timer value *)
   #at_tx[7] := #bit31;

   (* remember the last system time for the next overrun check *)
   #last_time := #tx;


   (* revision history
   DA  14.9.2007 rev 1.0
     original version

   DA  24.2.2008 rev 1.1
     added self reset on system startup

   DA   2.5.2008 rev 1.2
     corect a problem running under OB35

   DA  12.3.2009 rev 1.3
     corect a problem run on different CPUs

   DA  22.12.2009 rev 1.4
     corect a problem on startup
   *)
END_FUNCTION_BLOCK

FUNCTION_BLOCK "ALARM_2"   // FB122, SCL
TITLE = ALARM_2
{ S7_Optimized_Access := 'FALSE' }
AUTHOR : hugo
FAMILY : MEASURE
NAME : ALARM2
VERSION : 1.1
// ALARM_2 will check two pairs of limits and signal when the input is above or below a set limit.
// with the input HYS a hysteresis can be defined for all limits.
   VAR_INPUT
      X : Real;
      LO_1 : Real;
      HI_1 : Real;
      LO_2 : Real;
      HI_2 : Real;
      HYS : Real;
   END_VAR
   VAR_OUTPUT
      Q1_LO : Bool;
      Q1_HI : Bool;
      Q2_LO : Bool;
      Q2_HI : Bool;
   END_VAR
   VAR
      tmp : Real;
   END_VAR
BEGIN


   #tmp := #X - #HYS * 0.5;
   IF #tmp > #LO_1 THEN #Q1_LO := FALSE; END_IF;
   IF #tmp > #LO_2 THEN #Q2_LO := FALSE; END_IF;
   IF #tmp > #HI_1 THEN #Q1_HI := TRUE; END_IF;
   IF #tmp > #HI_2 THEN #Q2_HI := TRUE; END_IF;
   #tmp := #tmp + #HYS;
   IF #tmp < #LO_1 THEN #Q1_LO := TRUE; END_IF;
   IF #tmp < #LO_2 THEN #Q2_LO := TRUE; END_IF;
   IF #tmp < #HI_1 THEN #Q1_HI := FALSE; END_IF;
   IF #tmp < #HI_2 THEN #Q2_HI := FALSE; END_IF;


   (* revision history
   hm  19. may. 2008       rev 1.0
       original version

   hm  11. mar. 2009   rev 1.1
       improved code
   *)
END_FUNCTION_BLOCK

FUNCTION_BLOCK "BAR_GRAPH"   // FB123, SCL
TITLE = BAR_GRAPH
{ S7_Optimized_Access := 'FALSE' }
AUTHOR : hugo
FAMILY : MEASURE
NAME : BARGRAPH
VERSION : 1.2
// bar graph is a muti window comparator which displays an analog input signal on 8 digital outputs.
// only one output is active a any given time depending on the value of the input signal.
// the output can be of linear or logarithmic scale.
   VAR_INPUT
      X : Real;
      rst : Bool;
      trigger_Low : Real;
      trigger_High : Real;
      Alarm_low : Bool;
      Alarm_high : Bool;
      log_scale : Bool;
   END_VAR
   VAR_OUTPUT
      LOW : Bool;
      Q1 : Bool;
      Q2 : Bool;
      Q3 : Bool;
      Q4 : Bool;
      Q5 : Bool;
      Q6 : Bool;
      HIGH : Bool;
      Alarm : Bool;
      Status : Byte;
   END_VAR
   VAR
      init : Bool;
      T_1 : Real;
      T_2 : Real;
      T_3 : Real;
      T_4 : Real;
      T_5 : Real;
   END_VAR
   VAR_TEMP
      temp : Real;
   END_VAR
BEGIN


     IF NOT #init THEN
         #init := TRUE;
         IF #log_scale THEN
             #temp := (#trigger_High / #trigger_Low)**0.166666666666666666666;
             #T_1 := #trigger_Low * #temp;
             #T_2 := #T_1 * #temp;
             #T_3 := #T_2 * #temp;
             #T_4 := #T_3 * #temp;
             #T_5 := #T_4 * #temp;
         ELSE
             #temp := (#trigger_High - #trigger_Low) * 0.142857142;
             #T_1 := #trigger_Low + #temp;
             #T_2 := #T_1 + #temp;
             #T_3 := #T_2 + #temp;
             #T_4 := #T_3 + #temp;
             #T_5 := #T_4 + #temp;
         END_IF;
     END_IF;

   (* clear outputs before checking *)
     #Q1 := FALSE;
     #Q2 := FALSE;
     #Q3 := FALSE;
     #Q4 := FALSE;
     #Q5 := FALSE;
     #Q6 := FALSE;
     #Status := 110;

   (* low, high and alarm can only be cleared with rst depending on alarm_low and alarm_high *)
     IF NOT #Alarm_low THEN #LOW := FALSE; END_IF;
     IF NOT #Alarm_high THEN #HIGH := FALSE; END_IF;
     IF #rst THEN
         #Alarm := FALSE;
         #LOW := FALSE;
         #HIGH := FALSE;
     END_IF;

